(* Logix 5000 project; controller PLC_MCC1201_220AP1 vendor 1 type 14 code 164 rev 35.11; software revision 35.00; part 24 of 25 *)
(* tags used below, declared in another part *)
   dMaxLehrSpeed : DINT;
   dMinLehrSpeed : DINT;
   TMP_xDummy : BOOL;
   xAlwaysOFF : BOOL;
   N53 : DINT[10];
   N53_HOST : INT[10];
   N54 : DINT[501];
   TMP_xAlwaysOFF : BOOL;
   Z200 : MAC_Zone_ML;
   Z200_ALM : MAC_Zone_ML_ALM;
   Z200_HMR : MAC_Zone_ML_HMR;
   Z200_HMW : MAC_Zone_ML_HMW;
   Z200_UPS : ZONE_UPS;
   Z200_UPS_ALM : ZONE_UPS_ALM;
   Z200_UPS_HMR : ZONE_UPS_HMR;
   Z200_UPS_HMW : ZONE_UPS_HMW;
(* MainProgram, continued *)

ROUTINE Z200_Logics   (* ladder *)
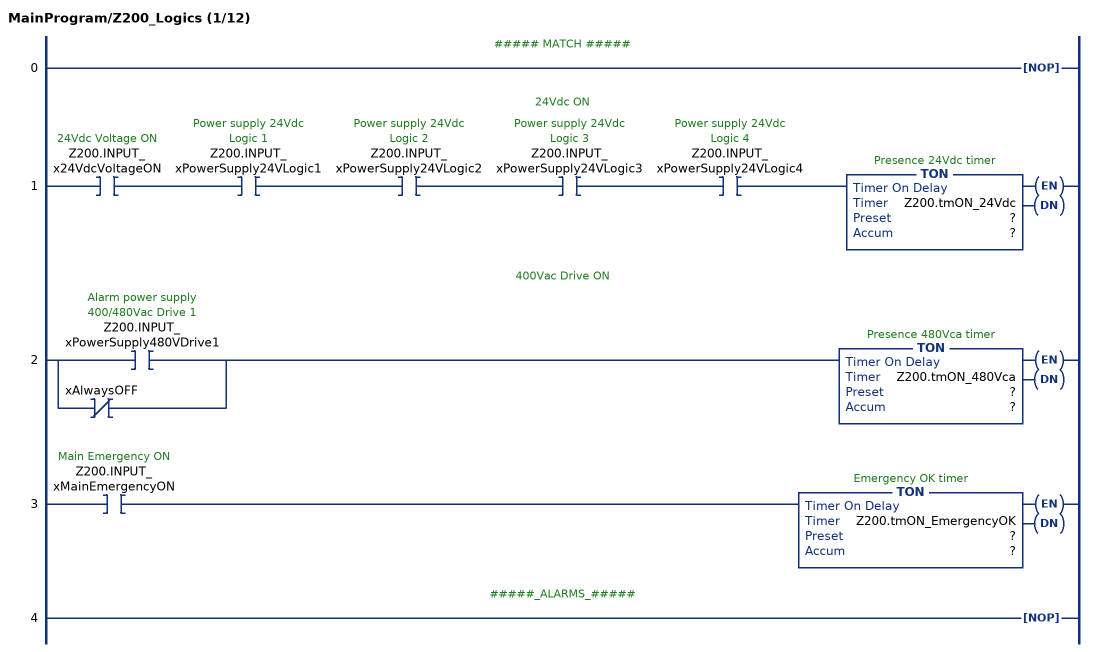
   // ##### MATCH #####
   0: NOP();
   // 24Vdc ON
   1: XIC(Z200.INPUT_x24VdcVoltageON)XIC(Z200.INPUT_xPowerSupply24VLogic1)XIC(Z200.INPUT_xPowerSupply24VLogic2)XIC(Z200.INPUT_xPowerSupply24VLogic3)XIC(Z200.INPUT_xPowerSupply24VLogic4)TON(Z200.tmON_24Vdc,?,?);
   // 400Vac Drive ON
   2: [XIC(Z200.INPUT_xPowerSupply480VDrive1) ,XIO(xAlwaysOFF) ]TON(Z200.tmON_480Vca,?,?);
   3: XIC(Z200.INPUT_xMainEmergencyON)TON(Z200.tmON_EmergencyOK,?,?);
   // #####_ALARMS_#####
   4: NOP();
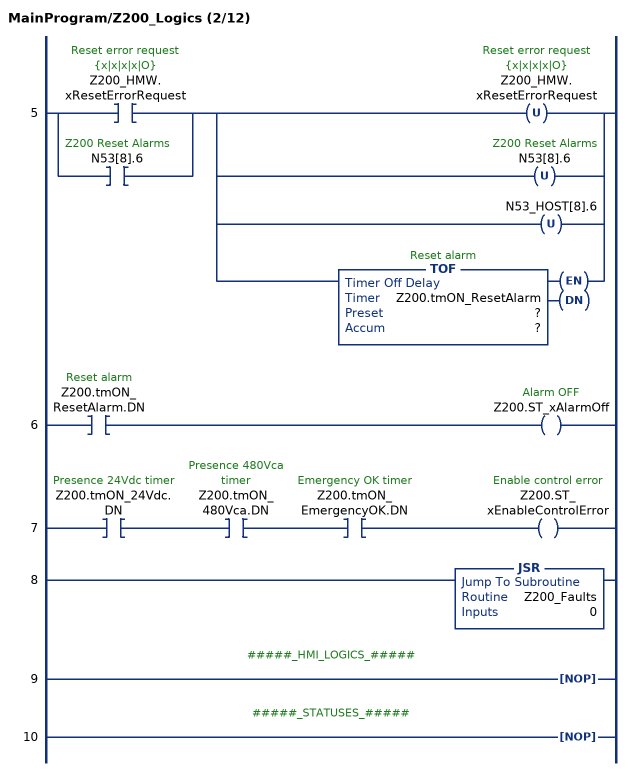
   5: [XIC(Z200_HMW.xResetErrorRequest) ,XIC(N53[8].6) ][OTU(Z200_HMW.xResetErrorRequest) ,OTU(N53[8].6) ,OTU(N53_HOST[8].6) ,TOF(Z200.tmON_ResetAlarm,?,?) ];
   6: XIC(Z200.tmON_ResetAlarm.DN)OTE(Z200.ST_xAlarmOff);
   7: XIC(Z200.tmON_24Vdc.DN)XIC(Z200.tmON_480Vca.DN)XIC(Z200.tmON_EmergencyOK.DN)OTE(Z200.ST_xEnableControlError);
   8: JSR(Z200_Faults,0);
   // #####_HMI_LOGICS_#####
   9: NOP();
   // #####_STATUSES_#####
   10: NOP();
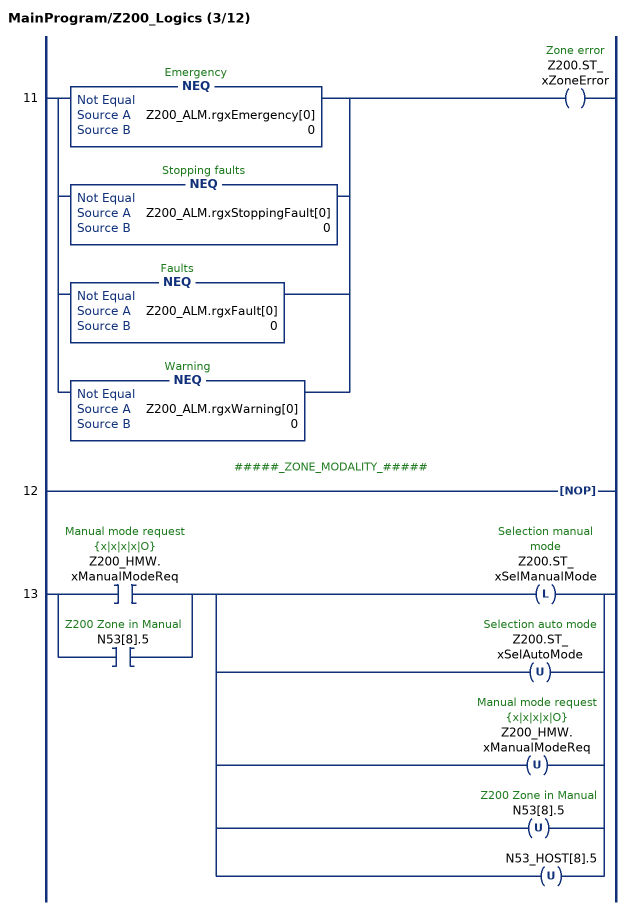
   11: [NEQ(Z200_ALM.rgxEmergency[0],0) ,NEQ(Z200_ALM.rgxStoppingFault[0],0) ,NEQ(Z200_ALM.rgxFault[0],0) ,NEQ(Z200_ALM.rgxWarning[0],0) ]OTE(Z200.ST_xZoneError);
   // #####_ZONE_MODALITY_#####
   12: NOP();
   13: [XIC(Z200_HMW.xManualModeReq) ,XIC(N53[8].5) ][OTL(Z200.ST_xSelManualMode) ,OTU(Z200.ST_xSelAutoMode) ,OTU(Z200_HMW.xManualModeReq) ,OTU(N53[8].5) ,OTU(N53_HOST[8].5) ];
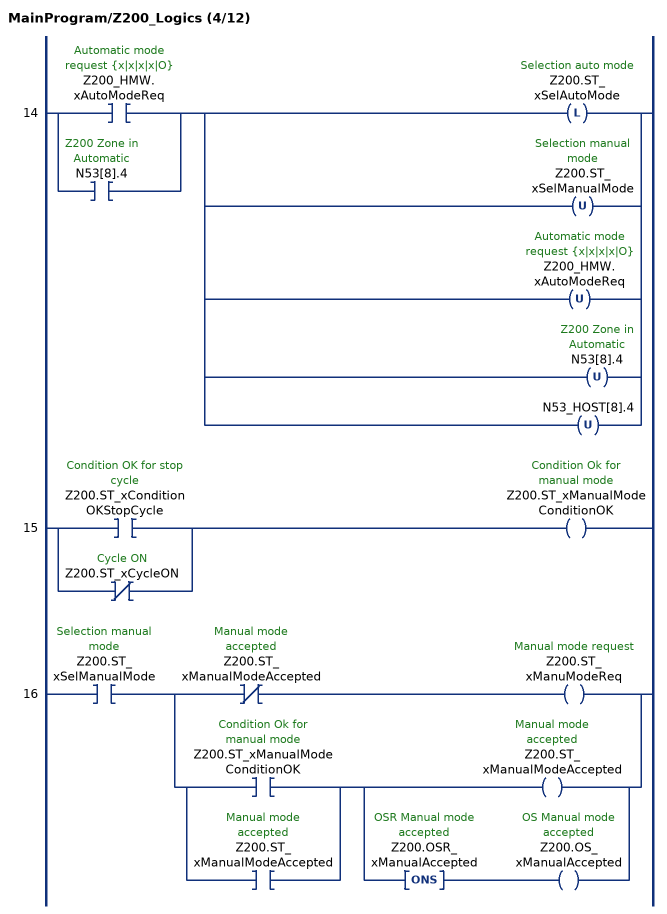
   14: [XIC(Z200_HMW.xAutoModeReq) ,XIC(N53[8].4) ][OTL(Z200.ST_xSelAutoMode) ,OTU(Z200.ST_xSelManualMode) ,OTU(Z200_HMW.xAutoModeReq) ,OTU(N53[8].4) ,OTU(N53_HOST[8].4) ];
   15: [XIC(Z200.ST_xConditionOKStopCycle) ,XIO(Z200.ST_xCycleON) ]OTE(Z200.ST_xManualModeConditionOK);
   16: XIC(Z200.ST_xSelManualMode)[XIO(Z200.ST_xManualModeAccepted) OTE(Z200.ST_xManuModeReq) ,[XIC(Z200.ST_xManualModeConditionOK) ,XIC(Z200.ST_xManualModeAccepted) ] [OTE(Z200.ST_xManualModeAccepted) ,ONS(Z200.OSR_xManualAccepted) OTE(Z200.OS_xManualAccepted) ] ];
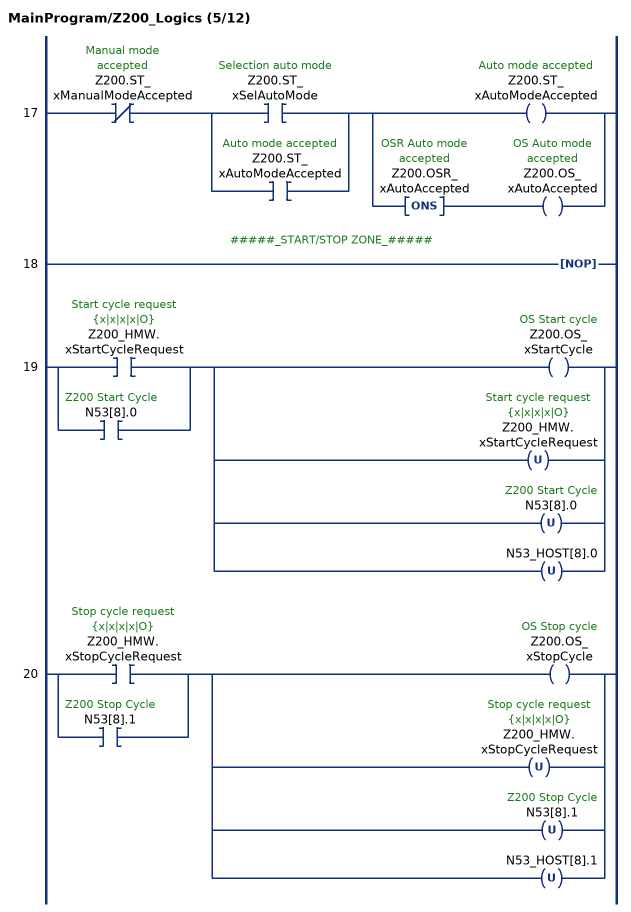
   17: XIO(Z200.ST_xManualModeAccepted)[XIC(Z200.ST_xSelAutoMode) ,XIC(Z200.ST_xAutoModeAccepted) ][OTE(Z200.ST_xAutoModeAccepted) ,ONS(Z200.OSR_xAutoAccepted) OTE(Z200.OS_xAutoAccepted) ];
   // #####_START/STOP ZONE_#####
   18: NOP();
   19: [XIC(Z200_HMW.xStartCycleRequest) ,XIC(N53[8].0) ][OTE(Z200.OS_xStartCycle) ,OTU(Z200_HMW.xStartCycleRequest) ,OTU(N53[8].0) ,OTU(N53_HOST[8].0) ];
   20: [XIC(Z200_HMW.xStopCycleRequest) ,XIC(N53[8].1) ][OTE(Z200.OS_xStopCycle) ,OTU(Z200_HMW.xStopCycleRequest) ,OTU(N53[8].1) ,OTU(N53_HOST[8].1) ];
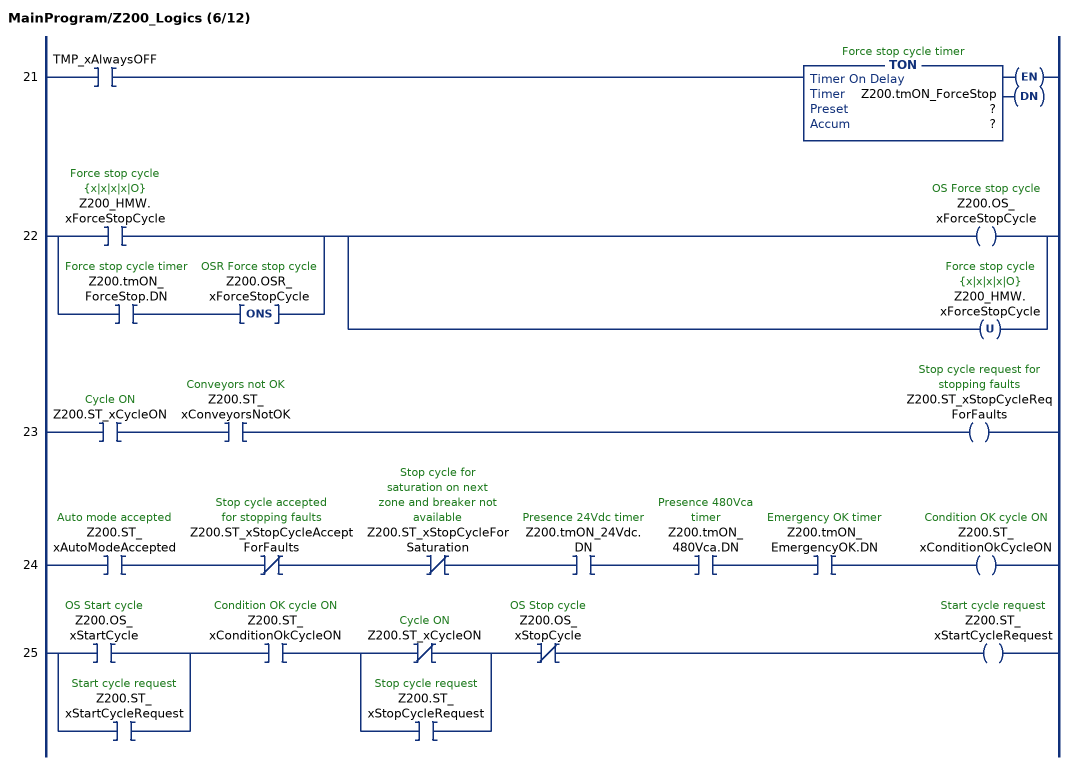
   21: XIC(TMP_xAlwaysOFF)TON(Z200.tmON_ForceStop,?,?);
   22: [XIC(Z200_HMW.xForceStopCycle) ,XIC(Z200.tmON_ForceStop.DN) ONS(Z200.OSR_xForceStopCycle) ][OTE(Z200.OS_xForceStopCycle) ,OTU(Z200_HMW.xForceStopCycle) ];
   23: XIC(Z200.ST_xCycleON)XIC(Z200.ST_xConveyorsNotOK)OTE(Z200.ST_xStopCycleReqForFaults);
   24: XIC(Z200.ST_xAutoModeAccepted)XIO(Z200.ST_xStopCycleAcceptForFaults)XIO(Z200.ST_xStopCycleForSaturation)XIC(Z200.tmON_24Vdc.DN)XIC(Z200.tmON_480Vca.DN)XIC(Z200.tmON_EmergencyOK.DN)OTE(Z200.ST_xConditionOkCycleON);
   25: [XIC(Z200.OS_xStartCycle) ,XIC(Z200.ST_xStartCycleRequest) ]XIC(Z200.ST_xConditionOkCycleON)[XIO(Z200.ST_xCycleON) ,XIC(Z200.ST_xStopCycleRequest) ]XIO(Z200.OS_xStopCycle)OTE(Z200.ST_xStartCycleRequest);
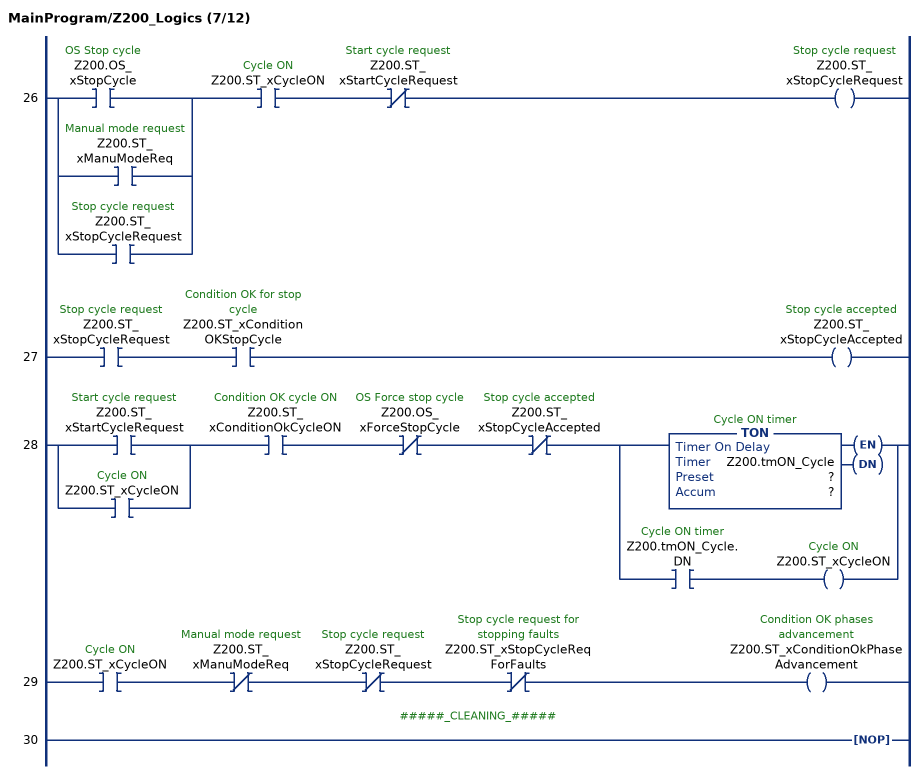
   26: [XIC(Z200.OS_xStopCycle) ,XIC(Z200.ST_xManuModeReq) ,XIC(Z200.ST_xStopCycleRequest) ]XIC(Z200.ST_xCycleON)XIO(Z200.ST_xStartCycleRequest)OTE(Z200.ST_xStopCycleRequest);
   27: XIC(Z200.ST_xStopCycleRequest)XIC(Z200.ST_xConditionOKStopCycle)OTE(Z200.ST_xStopCycleAccepted);
   28: [XIC(Z200.ST_xStartCycleRequest) ,XIC(Z200.ST_xCycleON) ]XIC(Z200.ST_xConditionOkCycleON)XIO(Z200.OS_xForceStopCycle)XIO(Z200.ST_xStopCycleAccepted)[TON(Z200.tmON_Cycle,?,?) ,XIC(Z200.tmON_Cycle.DN) OTE(Z200.ST_xCycleON) ];
   29: XIC(Z200.ST_xCycleON)XIO(Z200.ST_xManuModeReq)XIO(Z200.ST_xStopCycleRequest)XIO(Z200.ST_xStopCycleReqForFaults)OTE(Z200.ST_xConditionOkPhaseAdvancement);
   // #####_CLEANING_#####
   30: NOP();
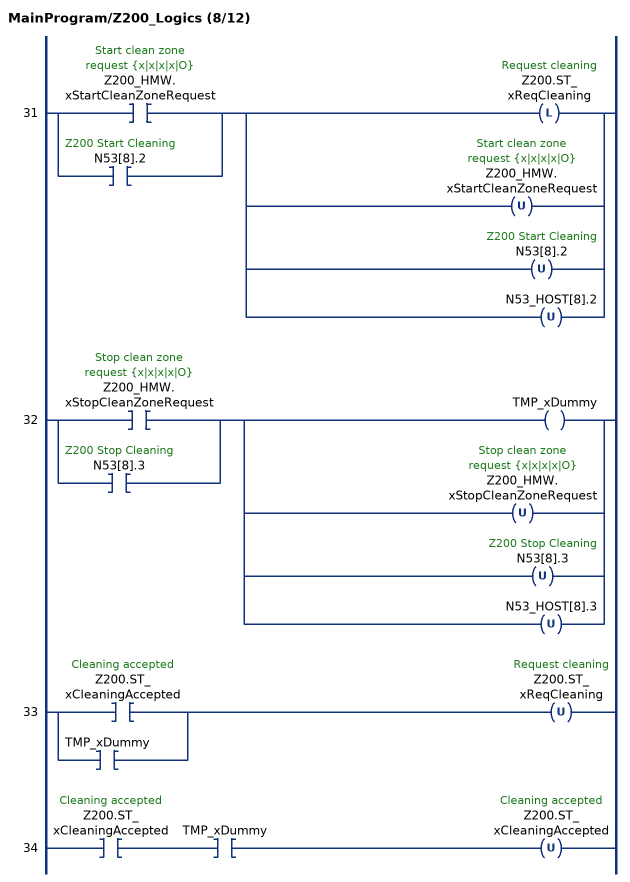
   31: [XIC(Z200_HMW.xStartCleanZoneRequest) ,XIC(N53[8].2) ][OTL(Z200.ST_xReqCleaning) ,OTU(Z200_HMW.xStartCleanZoneRequest) ,OTU(N53[8].2) ,OTU(N53_HOST[8].2) ];
   32: [XIC(Z200_HMW.xStopCleanZoneRequest) ,XIC(N53[8].3) ][OTE(TMP_xDummy) ,OTU(Z200_HMW.xStopCleanZoneRequest) ,OTU(N53[8].3) ,OTU(N53_HOST[8].3) ];
   33: [XIC(Z200.ST_xCleaningAccepted) ,XIC(TMP_xDummy) ]OTU(Z200.ST_xReqCleaning);
   34: XIC(Z200.ST_xCleaningAccepted)XIC(TMP_xDummy)OTU(Z200.ST_xCleaningAccepted);
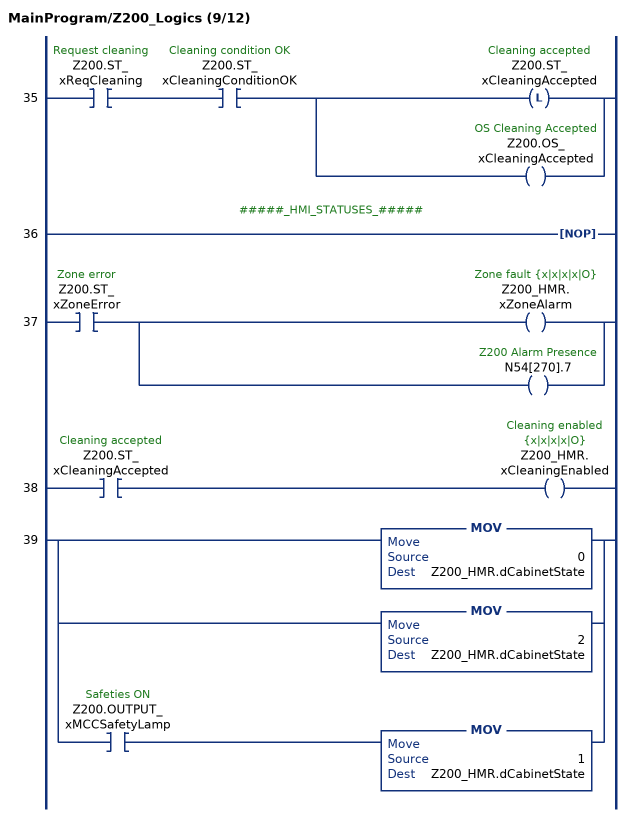
   35: XIC(Z200.ST_xReqCleaning)XIC(Z200.ST_xCleaningConditionOK)[OTL(Z200.ST_xCleaningAccepted) ,OTE(Z200.OS_xCleaningAccepted) ];
   // #####_HMI_STATUSES_#####
   36: NOP();
   37: XIC(Z200.ST_xZoneError)[OTE(Z200_HMR.xZoneAlarm) ,OTE(N54[270].7) ];
   38: XIC(Z200.ST_xCleaningAccepted)OTE(Z200_HMR.xCleaningEnabled);
   39: [MOV(0,Z200_HMR.dCabinetState) ,MOV(2,Z200_HMR.dCabinetState) ,XIC(Z200.OUTPUT_xMCCSafetyLamp) MOV(1,Z200_HMR.dCabinetState) ];
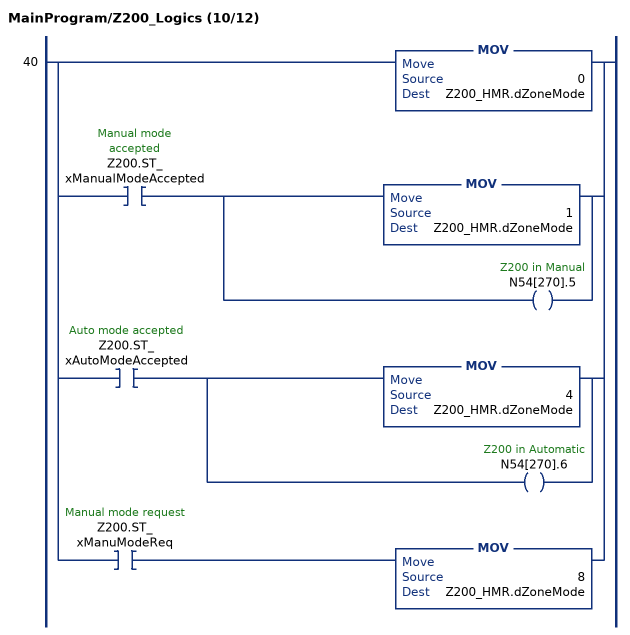
   40: [MOV(0,Z200_HMR.dZoneMode) ,XIC(Z200.ST_xManualModeAccepted) [MOV(1,Z200_HMR.dZoneMode) ,OTE(N54[270].5) ] ,XIC(Z200.ST_xAutoModeAccepted) [MOV(4,Z200_HMR.dZoneMode) ,OTE(N54[270].6) ] ,XIC(Z200.ST_xManuModeReq) MOV(8,Z200_HMR.dZoneMode) ];
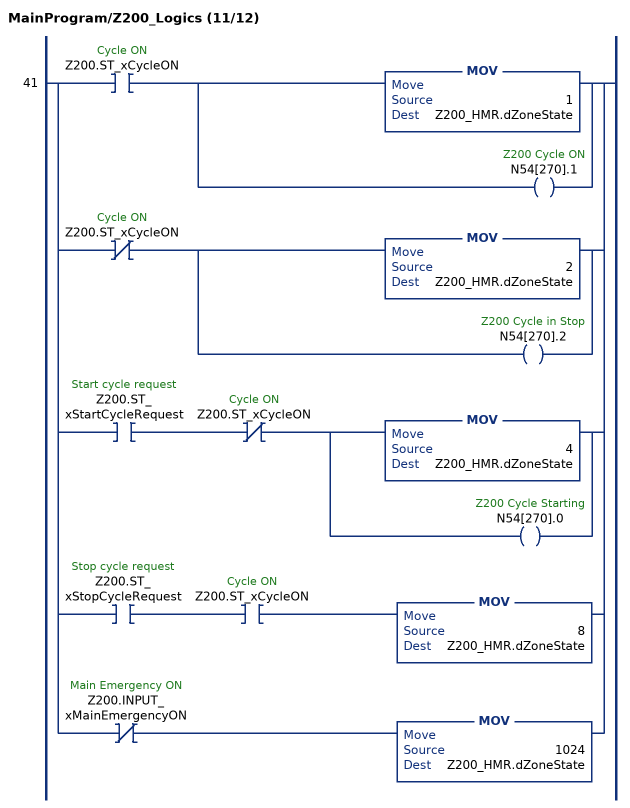
   41: [XIC(Z200.ST_xCycleON) [MOV(1,Z200_HMR.dZoneState) ,OTE(N54[270].1) ] ,XIO(Z200.ST_xCycleON) [MOV(2,Z200_HMR.dZoneState) ,OTE(N54[270].2) ] ,XIC(Z200.ST_xStartCycleRequest) XIO(Z200.ST_xCycleON) [MOV(4,Z200_HMR.dZoneState) ,OTE(N54[270].0) ] ,XIC(Z200.ST_xStopCycleRequest) XIC(Z200.ST_xCycleON) MOV(8,Z200_HMR.dZoneState) ,XIO(Z200.INPUT_xMainEmergencyON) MOV(1024,Z200_HMR.dZoneState) ];
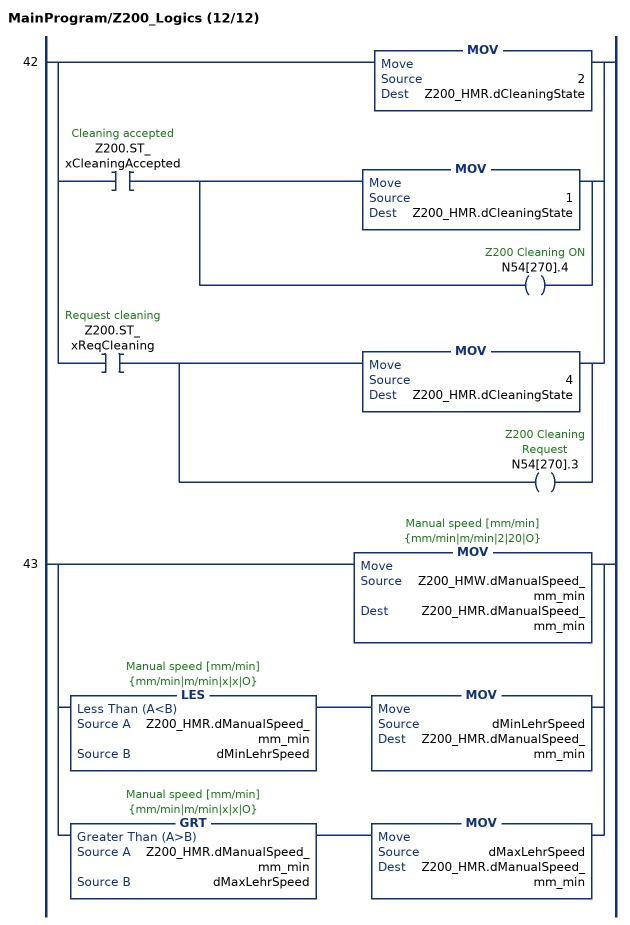
   42: [MOV(2,Z200_HMR.dCleaningState) ,XIC(Z200.ST_xCleaningAccepted) [MOV(1,Z200_HMR.dCleaningState) ,OTE(N54[270].4) ] ,XIC(Z200.ST_xReqCleaning) [MOV(4,Z200_HMR.dCleaningState) ,OTE(N54[270].3) ] ];
   43: [MOV(Z200_HMW.dManualSpeed_mm_min,Z200_HMR.dManualSpeed_mm_min) ,LES(Z200_HMR.dManualSpeed_mm_min,dMinLehrSpeed) MOV(dMinLehrSpeed,Z200_HMR.dManualSpeed_mm_min) ,GRT(Z200_HMR.dManualSpeed_mm_min,dMaxLehrSpeed) MOV(dMaxLehrSpeed,Z200_HMR.dManualSpeed_mm_min) ];
END_ROUTINE

ROUTINE Z200_UPS_Faults   (* ladder *)
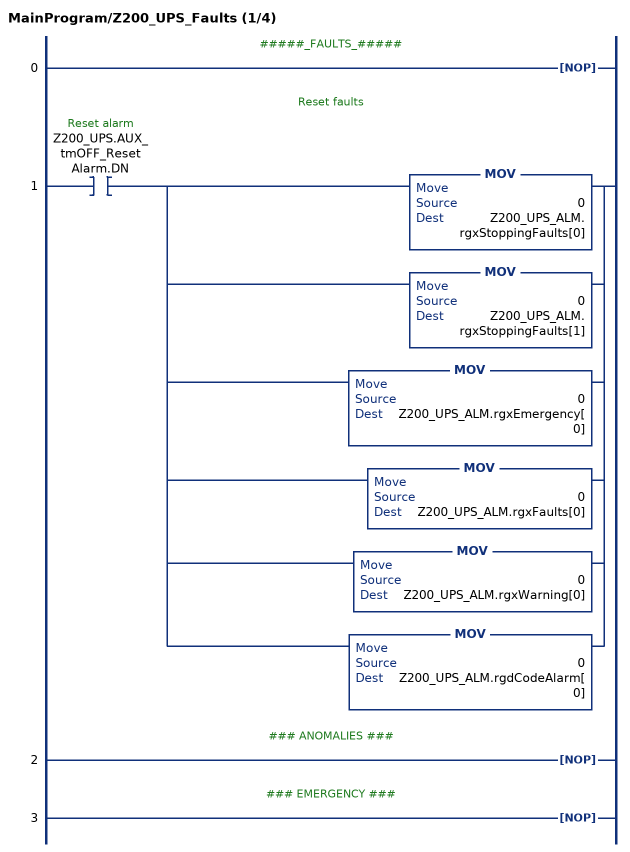
   // #####_FAULTS_#####
   0: NOP();
   // Reset faults
   1: XIC(Z200_UPS.AUX_tmOFF_ResetAlarm.DN)[MOV(0,Z200_UPS_ALM.rgxStoppingFaults[0]) ,MOV(0,Z200_UPS_ALM.rgxStoppingFaults[1]) ,MOV(0,Z200_UPS_ALM.rgxEmergency[0]) ,MOV(0,Z200_UPS_ALM.rgxFaults[0]) ,MOV(0,Z200_UPS_ALM.rgxWarning[0]) ,MOV(0,Z200_UPS_ALM.rgdCodeAlarm[0]) ];
   // ### ANOMALIES ###
   2: NOP();
   // ### EMERGENCY ###
   3: NOP();
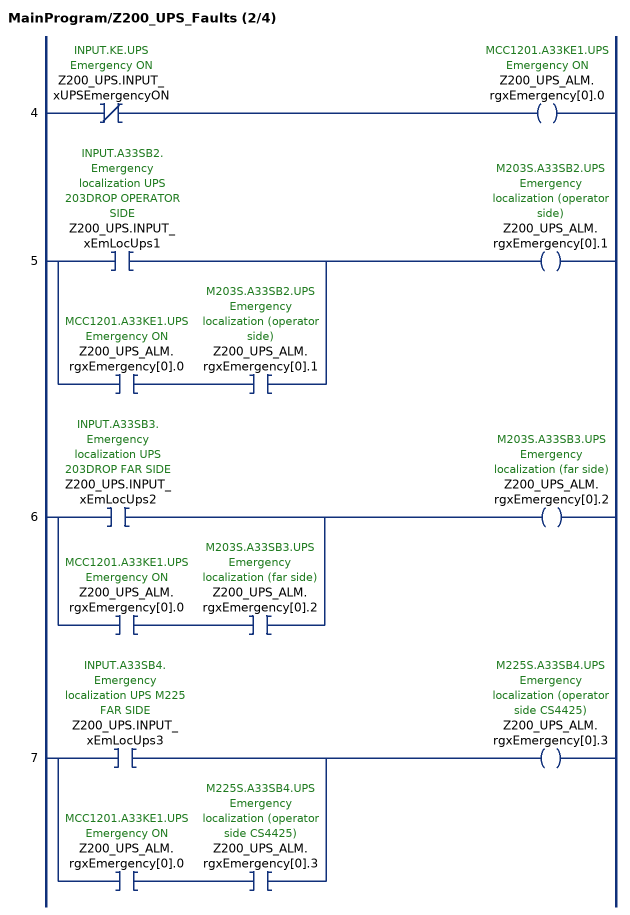
   4: XIO(Z200_UPS.INPUT_xUPSEmergencyON)OTE(Z200_UPS_ALM.rgxEmergency[0].0);
   5: [XIC(Z200_UPS.INPUT_xEmLocUps1) ,XIC(Z200_UPS_ALM.rgxEmergency[0].0) XIC(Z200_UPS_ALM.rgxEmergency[0].1) ]OTE(Z200_UPS_ALM.rgxEmergency[0].1);
   6: [XIC(Z200_UPS.INPUT_xEmLocUps2) ,XIC(Z200_UPS_ALM.rgxEmergency[0].0) XIC(Z200_UPS_ALM.rgxEmergency[0].2) ]OTE(Z200_UPS_ALM.rgxEmergency[0].2);
   7: [XIC(Z200_UPS.INPUT_xEmLocUps3) ,XIC(Z200_UPS_ALM.rgxEmergency[0].0) XIC(Z200_UPS_ALM.rgxEmergency[0].3) ]OTE(Z200_UPS_ALM.rgxEmergency[0].3);
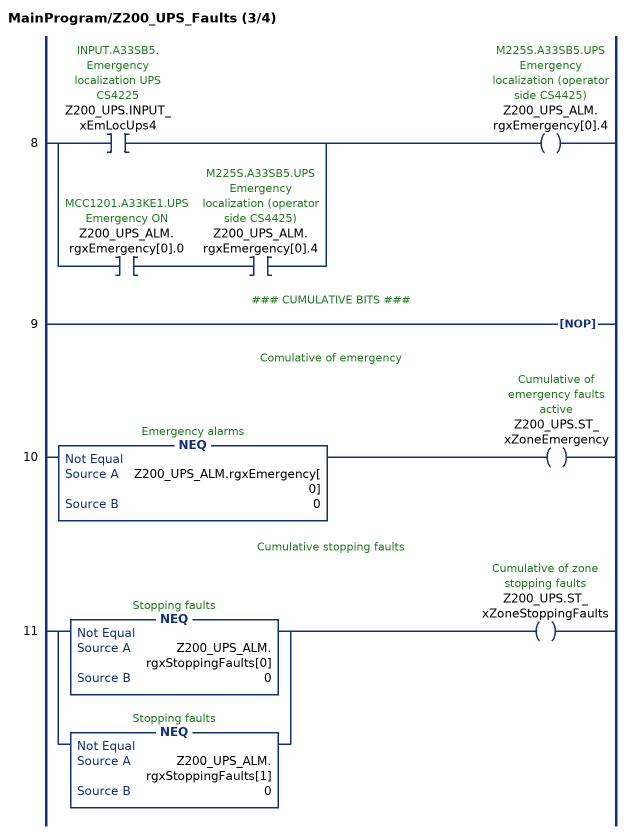
   8: [XIC(Z200_UPS.INPUT_xEmLocUps4) ,XIC(Z200_UPS_ALM.rgxEmergency[0].0) XIC(Z200_UPS_ALM.rgxEmergency[0].4) ]OTE(Z200_UPS_ALM.rgxEmergency[0].4);
   // ### CUMULATIVE BITS ###
   9: NOP();
   // Comulative of emergency
   10: NEQ(Z200_UPS_ALM.rgxEmergency[0],0)OTE(Z200_UPS.ST_xZoneEmergency);
   // Cumulative stopping faults
   11: [NEQ(Z200_UPS_ALM.rgxStoppingFaults[0],0) ,NEQ(Z200_UPS_ALM.rgxStoppingFaults[1],0) ]OTE(Z200_UPS.ST_xZoneStoppingFaults);
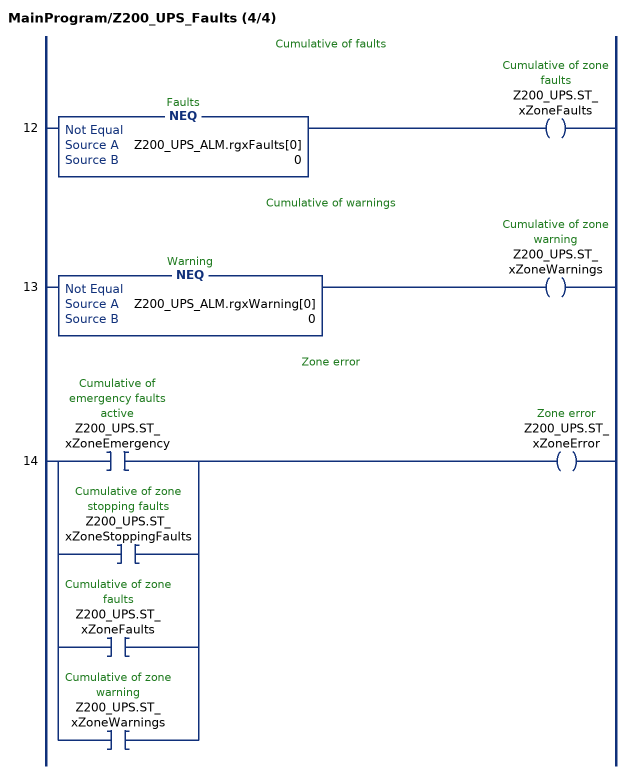
   // Cumulative of faults
   12: NEQ(Z200_UPS_ALM.rgxFaults[0],0)OTE(Z200_UPS.ST_xZoneFaults);
   // Cumulative of warnings
   13: NEQ(Z200_UPS_ALM.rgxWarning[0],0)OTE(Z200_UPS.ST_xZoneWarnings);
   // Zone error
   14: [XIC(Z200_UPS.ST_xZoneEmergency) ,XIC(Z200_UPS.ST_xZoneStoppingFaults) ,XIC(Z200_UPS.ST_xZoneFaults) ,XIC(Z200_UPS.ST_xZoneWarnings) ]OTE(Z200_UPS.ST_xZoneError);
END_ROUTINE

ROUTINE Z200_UPS_Logics   (* ladder *)
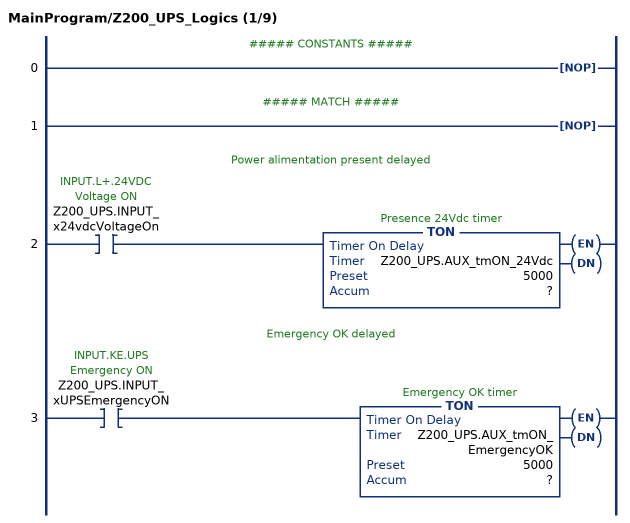
   // ##### CONSTANTS #####
   0: NOP();
   // ##### MATCH #####
   1: NOP();
   // Power alimentation present delayed
   2: XIC(Z200_UPS.INPUT_x24vdcVoltageOn)TON(Z200_UPS.AUX_tmON_24Vdc,?,?);
   // Emergency OK delayed
   3: XIC(Z200_UPS.INPUT_xUPSEmergencyON)TON(Z200_UPS.AUX_tmON_EmergencyOK,?,?);
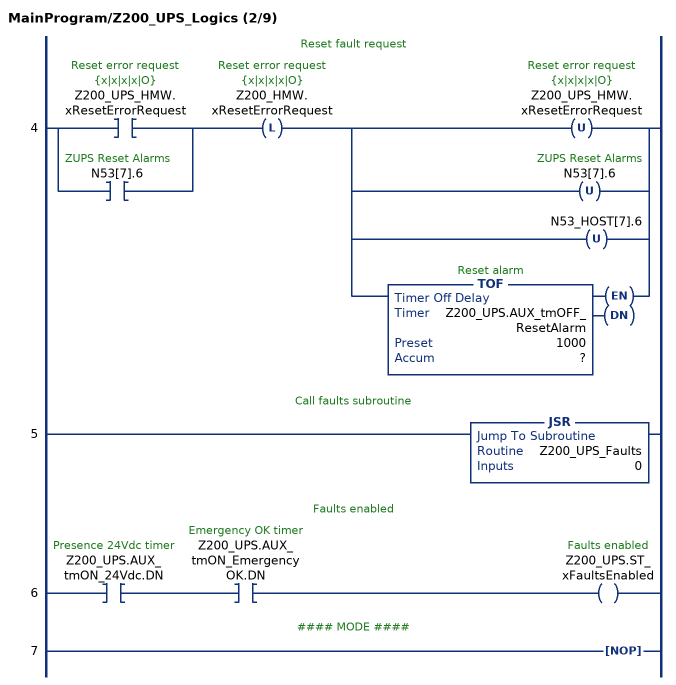
   // Reset fault request
   4: [XIC(Z200_UPS_HMW.xResetErrorRequest) ,XIC(N53[7].6) ]OTL(Z200_HMW.xResetErrorRequest)[OTU(Z200_UPS_HMW.xResetErrorRequest) ,OTU(N53[7].6) ,OTU(N53_HOST[7].6) ,TOF(Z200_UPS.AUX_tmOFF_ResetAlarm,?,?) ];
   // Call faults subroutine
   5: JSR(Z200_UPS_Faults,0);
   // Faults enabled
   6: XIC(Z200_UPS.AUX_tmON_24Vdc.DN)XIC(Z200_UPS.AUX_tmON_EmergencyOK.DN)OTE(Z200_UPS.ST_xFaultsEnabled);
   // #### MODE ####
   7: NOP();
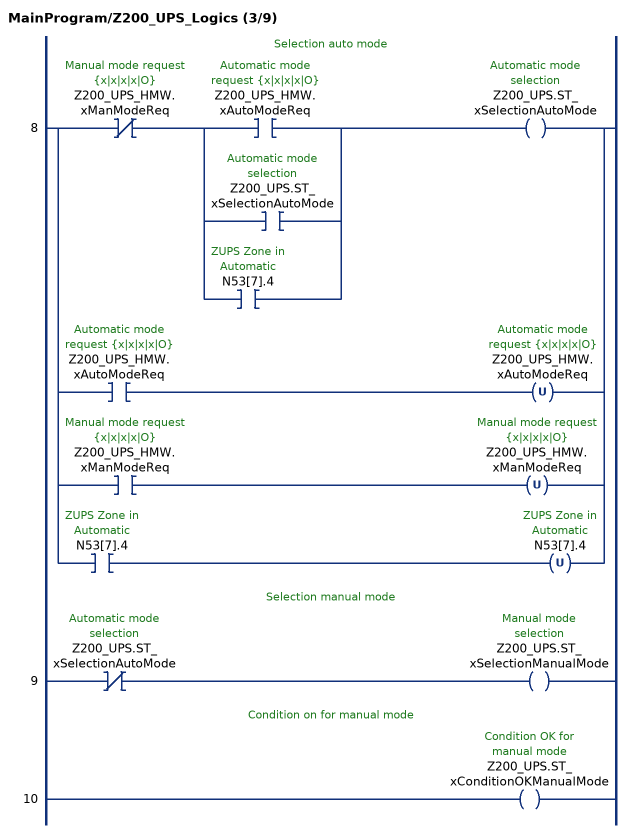
   // Selection auto mode
   8: [XIO(Z200_UPS_HMW.xManModeReq) [XIC(Z200_UPS_HMW.xAutoModeReq) ,XIC(Z200_UPS.ST_xSelectionAutoMode) ,XIC(N53[7].4) ] OTE(Z200_UPS.ST_xSelectionAutoMode) ,XIC(Z200_UPS_HMW.xAutoModeReq) OTU(Z200_UPS_HMW.xAutoModeReq) ,XIC(Z200_UPS_HMW.xManModeReq) OTU(Z200_UPS_HMW.xManModeReq) ,XIC(N53[7].4) OTU(N53[7].4) ];
   // Selection manual mode
   9: XIO(Z200_UPS.ST_xSelectionAutoMode)OTE(Z200_UPS.ST_xSelectionManualMode);
   // Condition on for manual mode
   10: OTE(Z200_UPS.ST_xConditionOKManualMode);
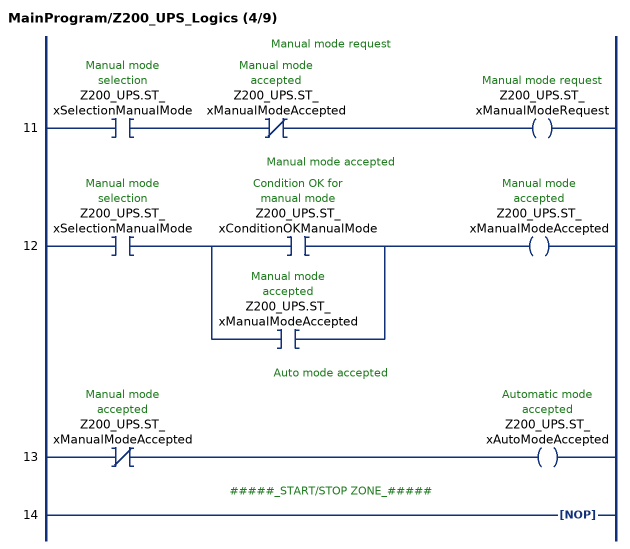
   // Manual mode request
   11: XIC(Z200_UPS.ST_xSelectionManualMode)XIO(Z200_UPS.ST_xManualModeAccepted)OTE(Z200_UPS.ST_xManualModeRequest);
   // Manual mode accepted
   12: XIC(Z200_UPS.ST_xSelectionManualMode)[XIC(Z200_UPS.ST_xConditionOKManualMode) ,XIC(Z200_UPS.ST_xManualModeAccepted) ]OTE(Z200_UPS.ST_xManualModeAccepted);
   // Auto mode accepted
   13: XIO(Z200_UPS.ST_xManualModeAccepted)OTE(Z200_UPS.ST_xAutoModeAccepted);
   // #####_START/STOP ZONE_#####
   14: NOP();
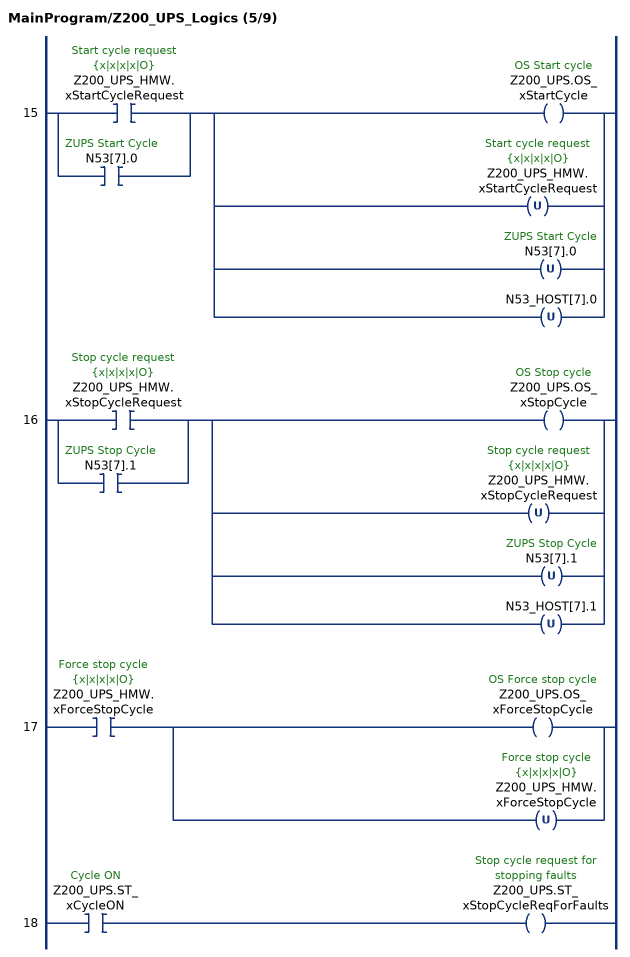
   15: [XIC(Z200_UPS_HMW.xStartCycleRequest) ,XIC(N53[7].0) ][OTE(Z200_UPS.OS_xStartCycle) ,OTU(Z200_UPS_HMW.xStartCycleRequest) ,OTU(N53[7].0) ,OTU(N53_HOST[7].0) ];
   16: [XIC(Z200_UPS_HMW.xStopCycleRequest) ,XIC(N53[7].1) ][OTE(Z200_UPS.OS_xStopCycle) ,OTU(Z200_UPS_HMW.xStopCycleRequest) ,OTU(N53[7].1) ,OTU(N53_HOST[7].1) ];
   17: XIC(Z200_UPS_HMW.xForceStopCycle)[OTE(Z200_UPS.OS_xForceStopCycle) ,OTU(Z200_UPS_HMW.xForceStopCycle) ];
   18: XIC(Z200_UPS.ST_xCycleON)OTE(Z200_UPS.ST_xStopCycleReqForFaults);
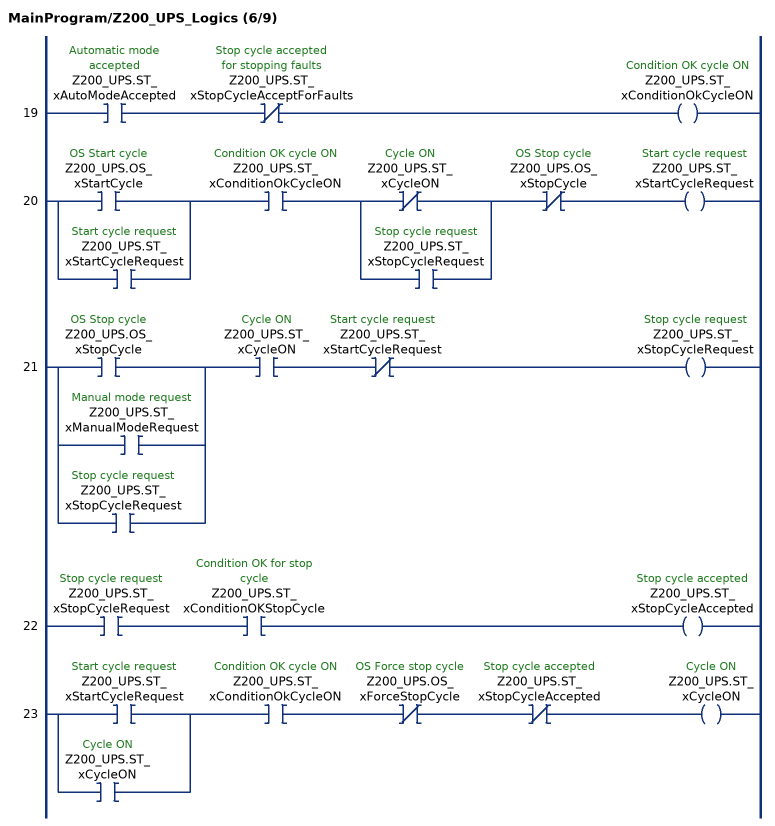
   19: XIC(Z200_UPS.ST_xAutoModeAccepted)XIO(Z200_UPS.ST_xStopCycleAcceptForFaults)OTE(Z200_UPS.ST_xConditionOkCycleON);
   20: [XIC(Z200_UPS.OS_xStartCycle) ,XIC(Z200_UPS.ST_xStartCycleRequest) ]XIC(Z200_UPS.ST_xConditionOkCycleON)[XIO(Z200_UPS.ST_xCycleON) ,XIC(Z200_UPS.ST_xStopCycleRequest) ]XIO(Z200_UPS.OS_xStopCycle)OTE(Z200_UPS.ST_xStartCycleRequest);
   21: [XIC(Z200_UPS.OS_xStopCycle) ,XIC(Z200_UPS.ST_xManualModeRequest) ,XIC(Z200_UPS.ST_xStopCycleRequest) ]XIC(Z200_UPS.ST_xCycleON)XIO(Z200_UPS.ST_xStartCycleRequest)OTE(Z200_UPS.ST_xStopCycleRequest);
   22: XIC(Z200_UPS.ST_xStopCycleRequest)XIC(Z200_UPS.ST_xConditionOKStopCycle)OTE(Z200_UPS.ST_xStopCycleAccepted);
   23: [XIC(Z200_UPS.ST_xStartCycleRequest) ,XIC(Z200_UPS.ST_xCycleON) ]XIC(Z200_UPS.ST_xConditionOkCycleON)XIO(Z200_UPS.OS_xForceStopCycle)XIO(Z200_UPS.ST_xStopCycleAccepted)OTE(Z200_UPS.ST_xCycleON);
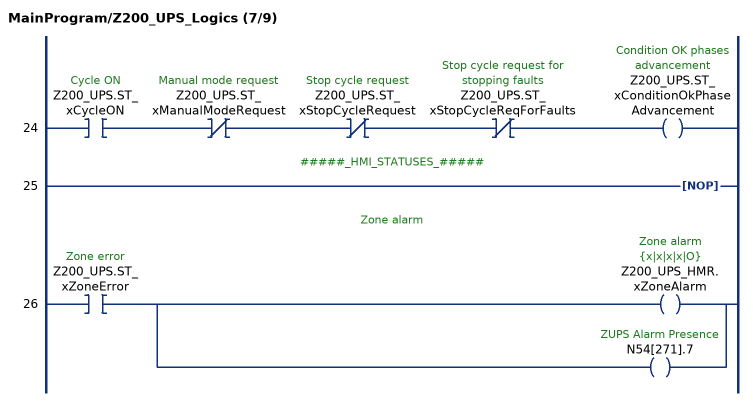
   24: XIC(Z200_UPS.ST_xCycleON)XIO(Z200_UPS.ST_xManualModeRequest)XIO(Z200_UPS.ST_xStopCycleRequest)XIO(Z200_UPS.ST_xStopCycleReqForFaults)OTE(Z200_UPS.ST_xConditionOkPhaseAdvancement);
   // #####_HMI_STATUSES_#####
   25: NOP();
   // Zone alarm
   26: XIC(Z200_UPS.ST_xZoneError)[OTE(Z200_UPS_HMR.xZoneAlarm) ,OTE(N54[271].7) ];
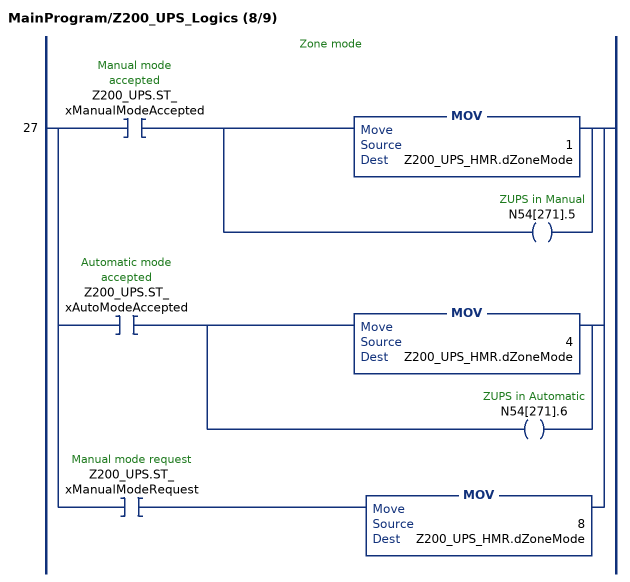
   // Zone mode
   27: [XIC(Z200_UPS.ST_xManualModeAccepted) [MOV(1,Z200_UPS_HMR.dZoneMode) ,OTE(N54[271].5) ] ,XIC(Z200_UPS.ST_xAutoModeAccepted) [MOV(4,Z200_UPS_HMR.dZoneMode) ,OTE(N54[271].6) ] ,XIC(Z200_UPS.ST_xManualModeRequest) MOV(8,Z200_UPS_HMR.dZoneMode) ];
